// TIA Portal project "消毒机" (V15.1) (continued)
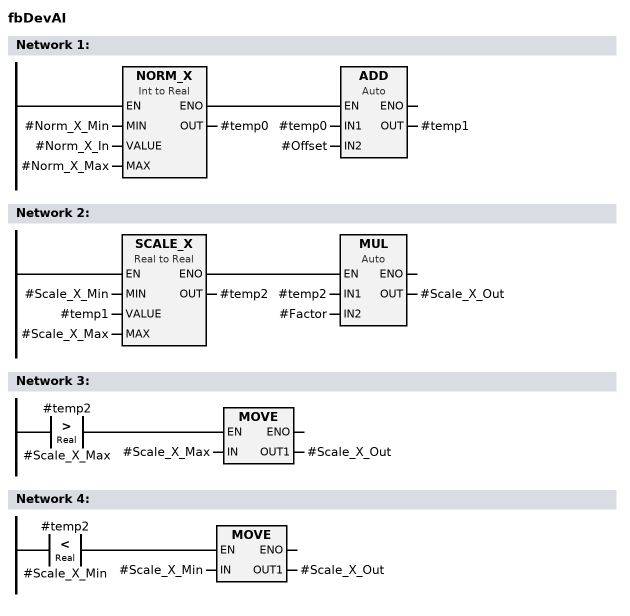
   RUNG wire#powerrail
      { S7_Templates := "[SrcType := Int, DestType := Real]" } Normalize(min := #Norm_X_Min, value := #Norm_X_In, max := #Norm_X_Max, out => #temp0)
      Add(in1 := #temp0, in2 := #Offset, out => #temp1)
   END_RUNG
   // the same network as SCL:
   #temp0 := NORM_X(MIN := #Norm_X_Min, VALUE := #Norm_X_In, MAX := #Norm_X_Max);
   #temp1 := #temp0 + #Offset;
END_REGION

REGION Network 2
   RUNG wire#powerrail
      { S7_Templates := "[SrcType := Real, DestType := Real]" } Scale(min := #Scale_X_Min, value := #temp1, max := #Scale_X_Max, out => #temp2)
      Mul(in1 := #temp2, in2 := #Factor, out => #Scale_X_Out)
   END_RUNG
   // the same network as SCL:
   #temp2 := SCALE_X(MIN := #Scale_X_Min, VALUE := #temp1, MAX := #Scale_X_Max);
   #Scale_X_Out := #temp2 * #Factor;
END_REGION

REGION Network 3
   RUNG wire#powerrail
      { S7_Templates := "SrcType := Real" } GT_Contact(in1 := #temp2, in2 := #Scale_X_Max)
      Move(in := #Scale_X_Max, out1 => #Scale_X_Out)
   END_RUNG
   // the same network as SCL:
   IF #temp2 > #Scale_X_Max THEN #Scale_X_Out := #Scale_X_Max; END_IF;
END_REGION

REGION Network 4
   RUNG wire#powerrail
      { S7_Templates := "SrcType := Real" } LT_Contact(in1 := #temp2, in2 := #Scale_X_Min)
      Move(in := #Scale_X_Min, out1 => #Scale_X_Out)
   END_RUNG
   // the same network as SCL:
   IF #temp2 < #Scale_X_Min THEN #Scale_X_Out := #Scale_X_Min; END_IF;
END_REGION
END_FUNCTION_BLOCK

FUNCTION_BLOCK "fbAI"   // FB102, LAD
{ S7_Optimized_Access := 'TRUE' }
VERSION : 0.1
   VAR
      fbDevAI_Instance : "fbDevAI";
      GET_IM_DATA_Instance : Get_IM_Data;
   END_VAR
   VAR_TEMP
      temp1 : Real;
   END_VAR
BEGIN

REGION Network 1
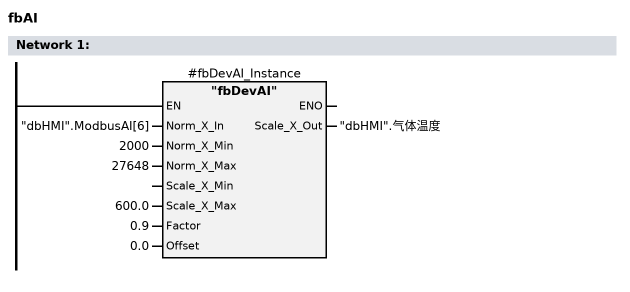
   RUNG wire#powerrail
      #fbDevAI_Instance(Norm_X_In := "dbHMI".ModbusAI[6], Norm_X_Min := 2000, Norm_X_Max := 27648, Scale_X_Min :=, Scale_X_Max := 600.0, Factor := 0.9, Offset := 0.0, Scale_X_Out => "dbHMI".气体温度)
   END_RUNG
   // the same network as SCL:
   #fbDevAI_Instance(Norm_X_In := "dbHMI".ModbusAI[6],   // "fbDevAI"
                     Norm_X_Min := 2000,
                     Norm_X_Max := 27648,
                     Scale_X_Max := 600.0,
                     Factor := 0.9,
                     Offset := 0.0,
                     Scale_X_Out => "dbHMI".气体温度);
END_REGION
END_FUNCTION_BLOCK

FUNCTION_BLOCK "fbSequence"   // FB103, LAD
{ S7_Optimized_Access := 'TRUE' }
VERSION : 0.1
   VAR_INPUT
      Start : Bool;
      Stop : Bool;
      ActUnit : "Unit";
   END_VAR
   VAR_OUTPUT
      ActStepNum : Int;
      OutUnit : "Unit";
   END_VAR
   VAR
      mRuntime_Step : Time;
      sRuntime_Step : Time;
      StepNo : Int;
      "Step" : Array[1..16] of Bool;
      StepDone : Array[1..16] of Bool;
      Next : Bool;
      StepStoped : Array[1..16] of Bool;
      Previos : Bool;
      IEC_Timer_1 : TON_TIME;
      IEC_Timer_2 : TON_TIME;
      IEC_Timer_3 : TON_TIME;
      IEC_Timer_4 : TON_TIME;
      IEC_Timer_5 : TON_TIME;
      IEC_Timer_6 : TON_TIME;
      IEC_Timer_7 : TON_TIME;
      IEC_Timer_8 : TON_TIME;
      IEC_Timer_9 : TON_TIME;
      IEC_Timer_10 : TON_TIME;
      IEC_Timer_11 : TON_TIME;
      IEC_Timer_12 : TON_TIME;
      IEC_Timer_13 : TON_TIME;
      IEC_Timer_14 : TON_TIME;
      IEC_Timer_15 : TON_TIME;
      IEC_Timer_16 : TON_TIME;
      Running : Bool;
      Done : Bool;
      Pls : Array[0..31] of Bool;
      AirCompressor_Step : Array[1..16] of Bool;
      Coolingwater_Step : Array[1..16] of Bool;
      Peristalticpump_Step : Array[1..16] of Bool;
      WepeX_Enable_Step : Array[1..16] of Bool;
      AYV1_Step : Array[1..16] of Bool;
      AYV2_Step : Array[1..16] of Bool;
      BYV1_Step : Array[1..16] of Bool;
      BYV2_Step : Array[1..16] of Bool;
      CYV1_Step : Array[1..16] of Bool;
      CYV2_Step : Array[1..16] of Bool;
      DYV_Step : Array[1..16] of Bool;
      Blower_Step : Array[1..16] of Bool;
   END_VAR
   VAR_TEMP   // added for the SCL form of the ladder/FBD networks
      _w1 : Bool;
   END_VAR
BEGIN

REGION Network 1
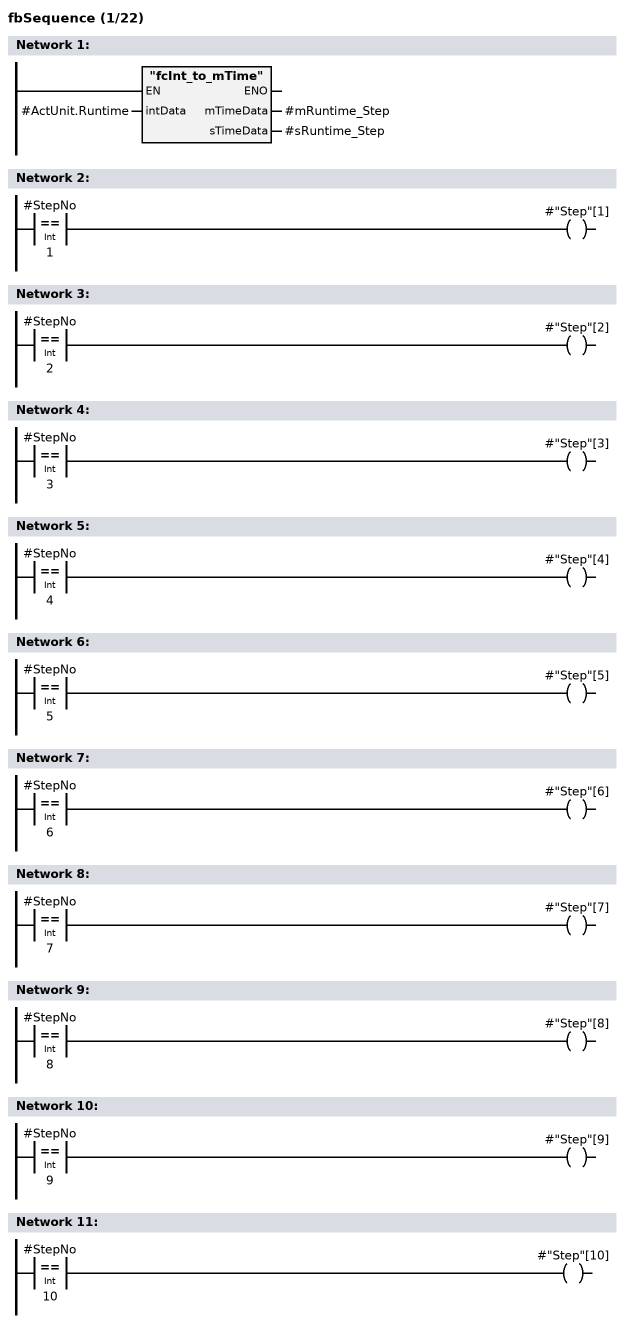
   RUNG wire#powerrail
      "fcInt_to_mTime"(intData := #ActUnit.Runtime, mTimeData => #mRuntime_Step, sTimeData => #sRuntime_Step)
   END_RUNG
   // the same network as SCL:
   "fcInt_to_mTime"(intData := #ActUnit.Runtime, mTimeData => #mRuntime_Step, sTimeData => #sRuntime_Step);
END_REGION

REGION Network 2
   RUNG wire#powerrail
      { S7_Templates := "SrcType := Int" } EQ_Contact(in1 := #StepNo, in2 := 1)
      Coil( #"Step"[1] )
   END_RUNG
   // the same network as SCL:
   #"Step"[1] := #StepNo = 1;
END_REGION

REGION Network 3
   RUNG wire#powerrail
      { S7_Templates := "SrcType := Int" } EQ_Contact(in1 := #StepNo, in2 := 2)
      Coil( #"Step"[2] )
   END_RUNG
   // the same network as SCL:
   #"Step"[2] := #StepNo = 2;
END_REGION

REGION Network 4
   RUNG wire#powerrail
      { S7_Templates := "SrcType := Int" } EQ_Contact(in1 := #StepNo, in2 := 3)
      Coil( #"Step"[3] )
   END_RUNG
   // the same network as SCL:
   #"Step"[3] := #StepNo = 3;
END_REGION

REGION Network 5
   RUNG wire#powerrail
      { S7_Templates := "SrcType := Int" } EQ_Contact(in1 := #StepNo, in2 := 4)
      Coil( #"Step"[4] )
   END_RUNG
   // the same network as SCL:
   #"Step"[4] := #StepNo = 4;
END_REGION

REGION Network 6
   RUNG wire#powerrail
      { S7_Templates := "SrcType := Int" } EQ_Contact(in1 := #StepNo, in2 := 5)
      Coil( #"Step"[5] )
   END_RUNG
   // the same network as SCL:
   #"Step"[5] := #StepNo = 5;
END_REGION

REGION Network 7
   RUNG wire#powerrail
      { S7_Templates := "SrcType := Int" } EQ_Contact(in1 := #StepNo, in2 := 6)
      Coil( #"Step"[6] )
   END_RUNG
   // the same network as SCL:
   #"Step"[6] := #StepNo = 6;
END_REGION

REGION Network 8
   RUNG wire#powerrail
      { S7_Templates := "SrcType := Int" } EQ_Contact(in1 := #StepNo, in2 := 7)
      Coil( #"Step"[7] )
   END_RUNG
   // the same network as SCL:
   #"Step"[7] := #StepNo = 7;
END_REGION

REGION Network 9
   RUNG wire#powerrail
      { S7_Templates := "SrcType := Int" } EQ_Contact(in1 := #StepNo, in2 := 8)
      Coil( #"Step"[8] )
   END_RUNG
   // the same network as SCL:
   #"Step"[8] := #StepNo = 8;
END_REGION

REGION Network 10
   RUNG wire#powerrail
      { S7_Templates := "SrcType := Int" } EQ_Contact(in1 := #StepNo, in2 := 9)
      Coil( #"Step"[9] )
   END_RUNG
   // the same network as SCL:
   #"Step"[9] := #StepNo = 9;
END_REGION

REGION Network 11
   RUNG wire#powerrail
      { S7_Templates := "SrcType := Int" } EQ_Contact(in1 := #StepNo, in2 := 10)
      Coil( #"Step"[10] )
   END_RUNG
   // the same network as SCL:
   #"Step"[10] := #StepNo = 10;
END_REGION

REGION Network 12
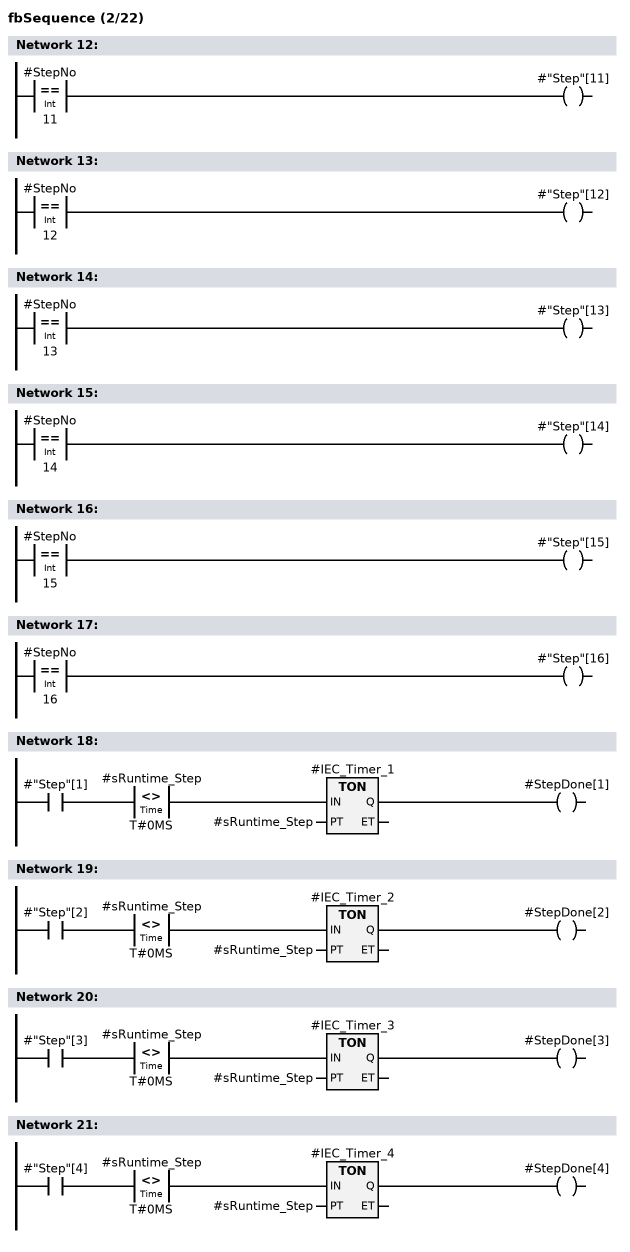
   RUNG wire#powerrail
      { S7_Templates := "SrcType := Int" } EQ_Contact(in1 := #StepNo, in2 := 11)
      Coil( #"Step"[11] )
   END_RUNG
   // the same network as SCL:
   #"Step"[11] := #StepNo = 11;
END_REGION

REGION Network 13
   RUNG wire#powerrail
      { S7_Templates := "SrcType := Int" } EQ_Contact(in1 := #StepNo, in2 := 12)
      Coil( #"Step"[12] )
   END_RUNG
   // the same network as SCL:
   #"Step"[12] := #StepNo = 12;
END_REGION

REGION Network 14
   RUNG wire#powerrail
      { S7_Templates := "SrcType := Int" } EQ_Contact(in1 := #StepNo, in2 := 13)
      Coil( #"Step"[13] )
   END_RUNG
   // the same network as SCL:
   #"Step"[13] := #StepNo = 13;
END_REGION

REGION Network 15
   RUNG wire#powerrail
      { S7_Templates := "SrcType := Int" } EQ_Contact(in1 := #StepNo, in2 := 14)
      Coil( #"Step"[14] )
   END_RUNG
   // the same network as SCL:
   #"Step"[14] := #StepNo = 14;
END_REGION

REGION Network 16
   RUNG wire#powerrail
      { S7_Templates := "SrcType := Int" } EQ_Contact(in1 := #StepNo, in2 := 15)
      Coil( #"Step"[15] )
   END_RUNG
   // the same network as SCL:
   #"Step"[15] := #StepNo = 15;
END_REGION

REGION Network 17
   RUNG wire#powerrail
      { S7_Templates := "SrcType := Int" } EQ_Contact(in1 := #StepNo, in2 := 16)
      Coil( #"Step"[16] )
   END_RUNG
   // the same network as SCL:
   #"Step"[16] := #StepNo = 16;
END_REGION

REGION Network 18
   #IEC_Timer_1(IN := #"Step"[1] AND (#sRuntime_Step <> T#0MS), PT := #sRuntime_Step);   // TON
   #StepDone[1] := #IEC_Timer_1.Q;
END_REGION

REGION Network 19
   #IEC_Timer_2(IN := #"Step"[2] AND (#sRuntime_Step <> T#0MS), PT := #sRuntime_Step);   // TON
   #StepDone[2] := #IEC_Timer_2.Q;
END_REGION

REGION Network 20
   #IEC_Timer_3(IN := #"Step"[3] AND (#sRuntime_Step <> T#0MS), PT := #sRuntime_Step);   // TON
   #StepDone[3] := #IEC_Timer_3.Q;
END_REGION

REGION Network 21
   #IEC_Timer_4(IN := #"Step"[4] AND (#sRuntime_Step <> T#0MS), PT := #sRuntime_Step);   // TON
   #StepDone[4] := #IEC_Timer_4.Q;
END_REGION

REGION Network 22
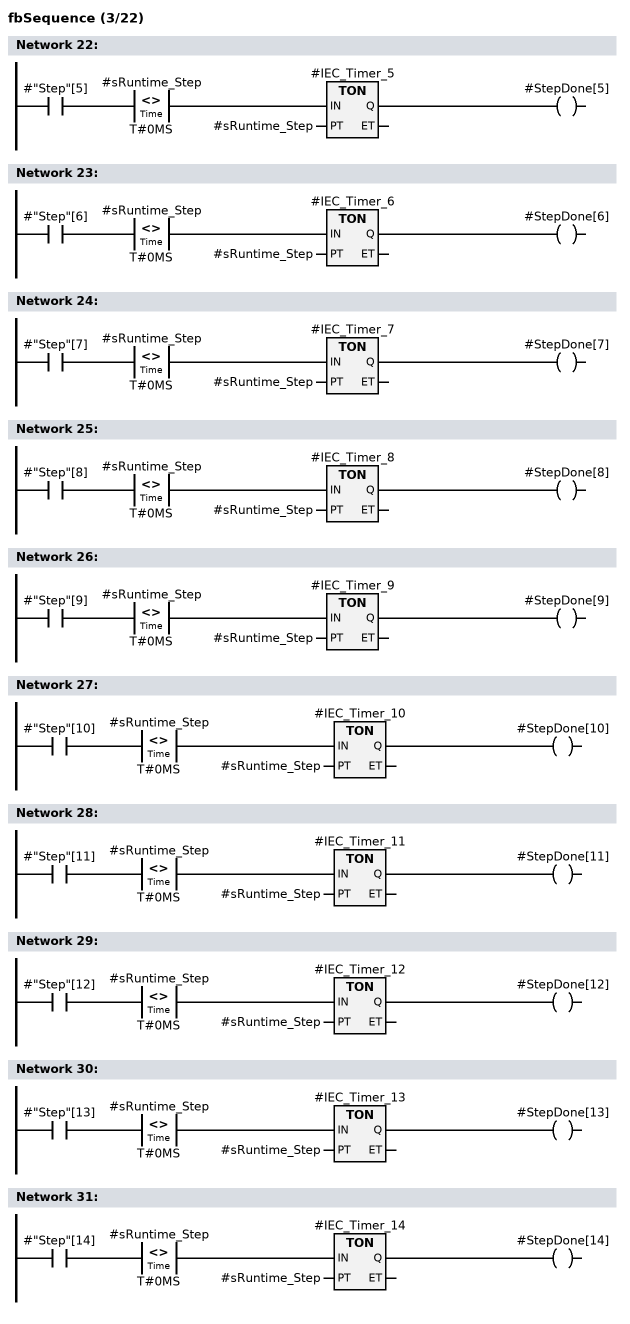
   #IEC_Timer_5(IN := #"Step"[5] AND (#sRuntime_Step <> T#0MS), PT := #sRuntime_Step);   // TON
   #StepDone[5] := #IEC_Timer_5.Q;
END_REGION

REGION Network 23
   #IEC_Timer_6(IN := #"Step"[6] AND (#sRuntime_Step <> T#0MS), PT := #sRuntime_Step);   // TON
   #StepDone[6] := #IEC_Timer_6.Q;
END_REGION

REGION Network 24
   #IEC_Timer_7(IN := #"Step"[7] AND (#sRuntime_Step <> T#0MS), PT := #sRuntime_Step);   // TON
   #StepDone[7] := #IEC_Timer_7.Q;
END_REGION

REGION Network 25
   #IEC_Timer_8(IN := #"Step"[8] AND (#sRuntime_Step <> T#0MS), PT := #sRuntime_Step);   // TON
   #StepDone[8] := #IEC_Timer_8.Q;
END_REGION

REGION Network 26
   #IEC_Timer_9(IN := #"Step"[9] AND (#sRuntime_Step <> T#0MS), PT := #sRuntime_Step);   // TON
   #StepDone[9] := #IEC_Timer_9.Q;
END_REGION

REGION Network 27
   #IEC_Timer_10(IN := #"Step"[10] AND (#sRuntime_Step <> T#0MS), PT := #sRuntime_Step);   // TON
   #StepDone[10] := #IEC_Timer_10.Q;
END_REGION

REGION Network 28
   #IEC_Timer_11(IN := #"Step"[11] AND (#sRuntime_Step <> T#0MS), PT := #sRuntime_Step);   // TON
   #StepDone[11] := #IEC_Timer_11.Q;
END_REGION

REGION Network 29
   #IEC_Timer_12(IN := #"Step"[12] AND (#sRuntime_Step <> T#0MS), PT := #sRuntime_Step);   // TON
   #StepDone[12] := #IEC_Timer_12.Q;
END_REGION

REGION Network 30
   #IEC_Timer_13(IN := #"Step"[13] AND (#sRuntime_Step <> T#0MS), PT := #sRuntime_Step);   // TON
   #StepDone[13] := #IEC_Timer_13.Q;
END_REGION

REGION Network 31
   #IEC_Timer_14(IN := #"Step"[14] AND (#sRuntime_Step <> T#0MS), PT := #sRuntime_Step);   // TON
   #StepDone[14] := #IEC_Timer_14.Q;
END_REGION

REGION Network 32
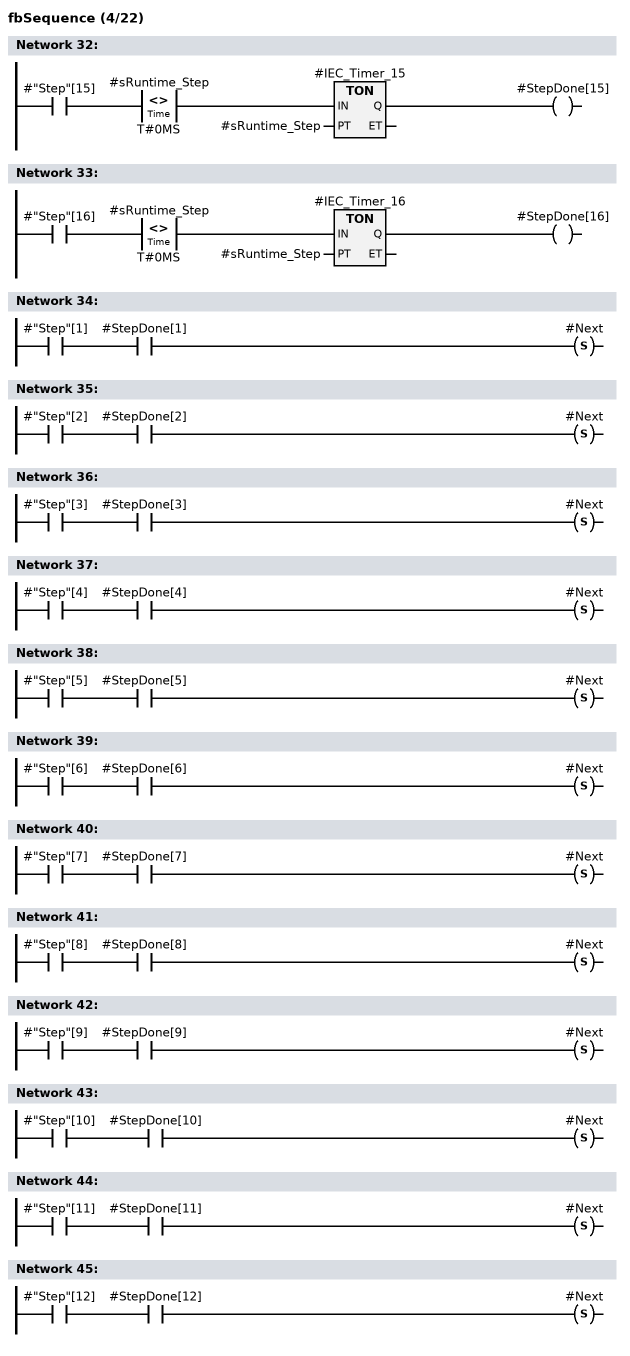
   #IEC_Timer_15(IN := #"Step"[15] AND (#sRuntime_Step <> T#0MS), PT := #sRuntime_Step);   // TON
   #StepDone[15] := #IEC_Timer_15.Q;
END_REGION

REGION Network 33
   #IEC_Timer_16(IN := #"Step"[16] AND (#sRuntime_Step <> T#0MS), PT := #sRuntime_Step);   // TON
   #StepDone[16] := #IEC_Timer_16.Q;
END_REGION

REGION Network 34
   RUNG wire#powerrail
      Contact( #"Step"[1] )
      Contact( #StepDone[1] )
      S_Coil( #Next )
   END_RUNG
   // the same network as SCL:
   IF #"Step"[1] AND #StepDone[1] THEN #Next := TRUE; END_IF;
END_REGION

REGION Network 35
   RUNG wire#powerrail
      Contact( #"Step"[2] )
      Contact( #StepDone[2] )
      S_Coil( #Next )
   END_RUNG
   // the same network as SCL:
   IF #"Step"[2] AND #StepDone[2] THEN #Next := TRUE; END_IF;
END_REGION

REGION Network 36
   RUNG wire#powerrail
      Contact( #"Step"[3] )
      Contact( #StepDone[3] )
      S_Coil( #Next )
   END_RUNG
   // the same network as SCL:
   IF #"Step"[3] AND #StepDone[3] THEN #Next := TRUE; END_IF;
END_REGION

REGION Network 37
   RUNG wire#powerrail
      Contact( #"Step"[4] )
      Contact( #StepDone[4] )
      S_Coil( #Next )
   END_RUNG
   // the same network as SCL:
   IF #"Step"[4] AND #StepDone[4] THEN #Next := TRUE; END_IF;
END_REGION

REGION Network 38
   RUNG wire#powerrail
      Contact( #"Step"[5] )
      Contact( #StepDone[5] )
      S_Coil( #Next )
   END_RUNG
   // the same network as SCL:
   IF #"Step"[5] AND #StepDone[5] THEN #Next := TRUE; END_IF;
END_REGION

REGION Network 39
   RUNG wire#powerrail
      Contact( #"Step"[6] )
      Contact( #StepDone[6] )
      S_Coil( #Next )
   END_RUNG
   // the same network as SCL:
   IF #"Step"[6] AND #StepDone[6] THEN #Next := TRUE; END_IF;
END_REGION

REGION Network 40
   RUNG wire#powerrail
      Contact( #"Step"[7] )
      Contact( #StepDone[7] )
      S_Coil( #Next )
   END_RUNG
   // the same network as SCL:
   IF #"Step"[7] AND #StepDone[7] THEN #Next := TRUE; END_IF;
END_REGION

REGION Network 41
   RUNG wire#powerrail
      Contact( #"Step"[8] )
      Contact( #StepDone[8] )
      S_Coil( #Next )
   END_RUNG
   // the same network as SCL:
   IF #"Step"[8] AND #StepDone[8] THEN #Next := TRUE; END_IF;
END_REGION

REGION Network 42
   RUNG wire#powerrail
      Contact( #"Step"[9] )
      Contact( #StepDone[9] )
      S_Coil( #Next )
   END_RUNG
   // the same network as SCL:
   IF #"Step"[9] AND #StepDone[9] THEN #Next := TRUE; END_IF;
END_REGION

REGION Network 43
   RUNG wire#powerrail
      Contact( #"Step"[10] )
      Contact( #StepDone[10] )
      S_Coil( #Next )
   END_RUNG
   // the same network as SCL:
   IF #"Step"[10] AND #StepDone[10] THEN #Next := TRUE; END_IF;
END_REGION

REGION Network 44
   RUNG wire#powerrail
      Contact( #"Step"[11] )
      Contact( #StepDone[11] )
      S_Coil( #Next )
   END_RUNG
   // the same network as SCL:
   IF #"Step"[11] AND #StepDone[11] THEN #Next := TRUE; END_IF;
END_REGION

REGION Network 45
   RUNG wire#powerrail
      Contact( #"Step"[12] )
      Contact( #StepDone[12] )
      S_Coil( #Next )
   END_RUNG
   // the same network as SCL:
   IF #"Step"[12] AND #StepDone[12] THEN #Next := TRUE; END_IF;
END_REGION

REGION Network 46
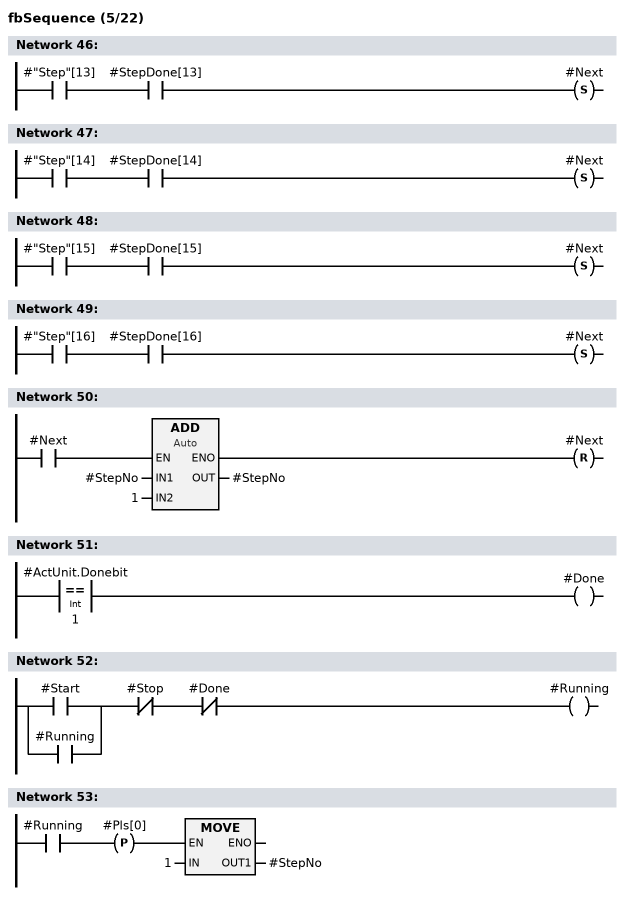
   RUNG wire#powerrail
      Contact( #"Step"[13] )
      Contact( #StepDone[13] )
      S_Coil( #Next )
   END_RUNG
   // the same network as SCL:
   IF #"Step"[13] AND #StepDone[13] THEN #Next := TRUE; END_IF;
END_REGION

REGION Network 47
   RUNG wire#powerrail
      Contact( #"Step"[14] )
      Contact( #StepDone[14] )
      S_Coil( #Next )
   END_RUNG
   // the same network as SCL:
   IF #"Step"[14] AND #StepDone[14] THEN #Next := TRUE; END_IF;
END_REGION

REGION Network 48
   RUNG wire#powerrail
      Contact( #"Step"[15] )
      Contact( #StepDone[15] )
      S_Coil( #Next )
   END_RUNG
   // the same network as SCL:
   IF #"Step"[15] AND #StepDone[15] THEN #Next := TRUE; END_IF;
END_REGION

REGION Network 49
   RUNG wire#powerrail
      Contact( #"Step"[16] )
      Contact( #StepDone[16] )
      S_Coil( #Next )
   END_RUNG
   // the same network as SCL:
   IF #"Step"[16] AND #StepDone[16] THEN #Next := TRUE; END_IF;
END_REGION

REGION Network 50
   RUNG wire#powerrail
      Contact( #Next )
      Add(in1 := #StepNo, in2 := 1, out => #StepNo)
      R_Coil( #Next )
   END_RUNG
   // the same network as SCL:
   IF #Next THEN
       #StepNo := #StepNo + 1;
       #Next := FALSE;
   END_IF;
END_REGION

REGION Network 51
   RUNG wire#powerrail
      { S7_Templates := "SrcType := Int" } EQ_Contact(in1 := #ActUnit.Donebit, in2 := 1)
      Coil( #Done )
   END_RUNG
   // the same network as SCL:
   #Done := #ActUnit.Donebit = 1;
END_REGION

REGION Network 52
   RUNG wire#powerrail
      Contact( #Start )
      wire#w1
      I_Contact( #Stop )
      I_Contact( #Done )
      Coil( #Running )
   END_RUNG
   RUNG wire#powerrail
      Contact( #Running )
   END_RUNG wire#w1
   // the same network as SCL:
   #Running := (#Start OR #Running) AND NOT #Stop AND NOT #Done;
END_REGION

REGION Network 53
   RUNG wire#powerrail
      Contact( #Running )
      P_Trig( #Pls[0] )
      Move(in := 1, out1 => #StepNo)
   END_RUNG
   // the same network as SCL:
   #_w1 := #Running AND NOT #Pls[0];   // rising edge
   #Pls[0] := #Running;
   IF #_w1 THEN #StepNo := 1; END_IF;
END_REGION

REGION Network 54
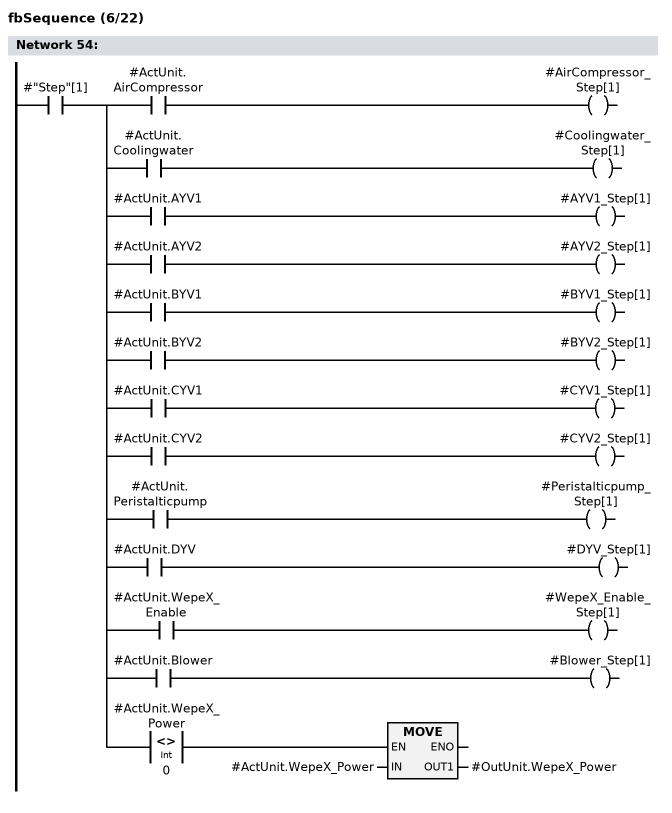
   RUNG wire#powerrail
      Contact( #"Step"[1] )
      wire#w1
      Contact( #ActUnit.AirCompressor )
      Coil( #AirCompressor_Step[1] )
   END_RUNG
   RUNG wire#w1
      Contact( #ActUnit.Coolingwater )
      Coil( #Coolingwater_Step[1] )
   END_RUNG
   RUNG wire#w1
      Contact( #ActUnit.AYV1 )
      Coil( #AYV1_Step[1] )
   END_RUNG
   RUNG wire#w1
      Contact( #ActUnit.AYV2 )
      Coil( #AYV2_Step[1] )
   END_RUNG
   RUNG wire#w1
      Contact( #ActUnit.BYV1 )
      Coil( #BYV1_Step[1] )
   END_RUNG
   RUNG wire#w1
      Contact( #ActUnit.BYV2 )
      Coil( #BYV2_Step[1] )
   END_RUNG
   RUNG wire#w1
      Contact( #ActUnit.CYV1 )
      Coil( #CYV1_Step[1] )
   END_RUNG
   RUNG wire#w1
      Contact( #ActUnit.CYV2 )
      Coil( #CYV2_Step[1] )
   END_RUNG
   RUNG wire#w1
      Contact( #ActUnit.Peristalticpump )
      Coil( #Peristalticpump_Step[1] )
   END_RUNG
   RUNG wire#w1
      Contact( #ActUnit.DYV )
      Coil( #DYV_Step[1] )
   END_RUNG
   RUNG wire#w1
      Contact( #ActUnit.WepeX_Enable )
      Coil( #WepeX_Enable_Step[1] )
   END_RUNG
   RUNG wire#w1
      Contact( #ActUnit.Blower )
      Coil( #Blower_Step[1] )
   END_RUNG
   RUNG wire#w1
      { S7_Templates := "SrcType := Int" } NE_Contact(in1 := #ActUnit.WepeX_Power, in2 := 0)
      Move(in := #ActUnit.WepeX_Power, out1 => #OutUnit.WepeX_Power)
   END_RUNG
   // the same network as SCL:
   #AirCompressor_Step[1] := #"Step"[1] AND #ActUnit.AirCompressor;
   #Coolingwater_Step[1] := #"Step"[1] AND #ActUnit.Coolingwater;
   #AYV1_Step[1] := #"Step"[1] AND #ActUnit.AYV1;
   #AYV2_Step[1] := #"Step"[1] AND #ActUnit.AYV2;
   #BYV1_Step[1] := #"Step"[1] AND #ActUnit.BYV1;
   #BYV2_Step[1] := #"Step"[1] AND #ActUnit.BYV2;
   #CYV1_Step[1] := #"Step"[1] AND #ActUnit.CYV1;
   #CYV2_Step[1] := #"Step"[1] AND #ActUnit.CYV2;
   #Peristalticpump_Step[1] := #"Step"[1] AND #ActUnit.Peristalticpump;
   #DYV_Step[1] := #"Step"[1] AND #ActUnit.DYV;
   #WepeX_Enable_Step[1] := #"Step"[1] AND #ActUnit.WepeX_Enable;
   #Blower_Step[1] := #"Step"[1] AND #ActUnit.Blower;
   IF #"Step"[1] AND (#ActUnit.WepeX_Power <> 0) THEN #OutUnit.WepeX_Power := #ActUnit.WepeX_Power; END_IF;
END_REGION

REGION Network 55
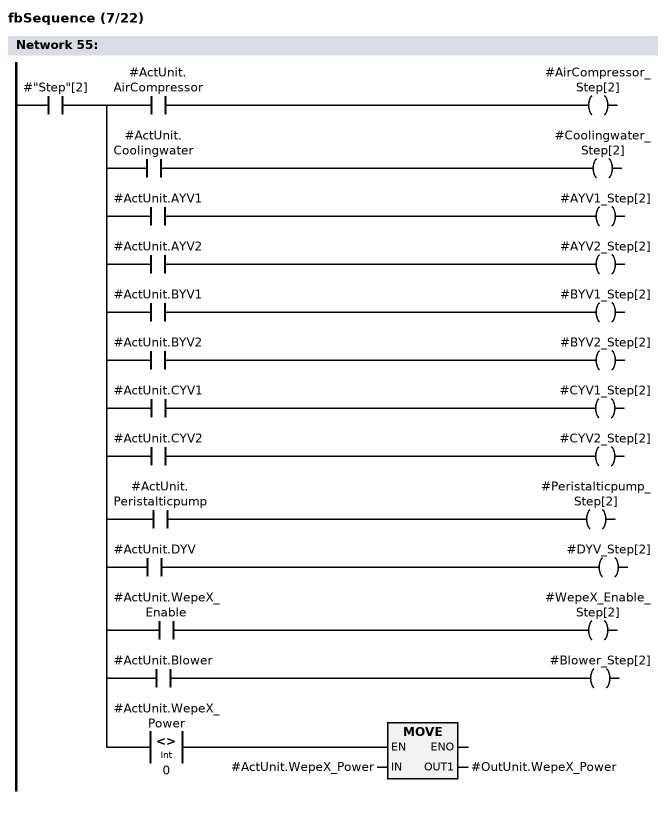
   RUNG wire#powerrail
      Contact( #"Step"[2] )
      wire#w1
      Contact( #ActUnit.AirCompressor )
      Coil( #AirCompressor_Step[2] )
   END_RUNG
   RUNG wire#w1
      Contact( #ActUnit.Coolingwater )
      Coil( #Coolingwater_Step[2] )
   END_RUNG
   RUNG wire#w1
      Contact( #ActUnit.AYV1 )
      Coil( #AYV1_Step[2] )
   END_RUNG
   RUNG wire#w1
      Contact( #ActUnit.AYV2 )
      Coil( #AYV2_Step[2] )
   END_RUNG
   RUNG wire#w1
      Contact( #ActUnit.BYV1 )
      Coil( #BYV1_Step[2] )
   END_RUNG
   RUNG wire#w1
      Contact( #ActUnit.BYV2 )
      Coil( #BYV2_Step[2] )
   END_RUNG
   RUNG wire#w1
      Contact( #ActUnit.CYV1 )
      Coil( #CYV1_Step[2] )
   END_RUNG
   RUNG wire#w1
      Contact( #ActUnit.CYV2 )
      Coil( #CYV2_Step[2] )
   END_RUNG
   RUNG wire#w1
      Contact( #ActUnit.Peristalticpump )
      Coil( #Peristalticpump_Step[2] )
   END_RUNG
   RUNG wire#w1
      Contact( #ActUnit.DYV )
      Coil( #DYV_Step[2] )
   END_RUNG
   RUNG wire#w1
      Contact( #ActUnit.WepeX_Enable )
      Coil( #WepeX_Enable_Step[2] )
   END_RUNG
   RUNG wire#w1
      Contact( #ActUnit.Blower )
      Coil( #Blower_Step[2] )
   END_RUNG
   RUNG wire#w1
      { S7_Templates := "SrcType := Int" } NE_Contact(in1 := #ActUnit.WepeX_Power, in2 := 0)
      Move(in := #ActUnit.WepeX_Power, out1 => #OutUnit.WepeX_Power)
   END_RUNG
   // the same network as SCL:
   #AirCompressor_Step[2] := #"Step"[2] AND #ActUnit.AirCompressor;
   #Coolingwater_Step[2] := #"Step"[2] AND #ActUnit.Coolingwater;
   #AYV1_Step[2] := #"Step"[2] AND #ActUnit.AYV1;
   #AYV2_Step[2] := #"Step"[2] AND #ActUnit.AYV2;
   #BYV1_Step[2] := #"Step"[2] AND #ActUnit.BYV1;
   #BYV2_Step[2] := #"Step"[2] AND #ActUnit.BYV2;
   #CYV1_Step[2] := #"Step"[2] AND #ActUnit.CYV1;
   #CYV2_Step[2] := #"Step"[2] AND #ActUnit.CYV2;
   #Peristalticpump_Step[2] := #"Step"[2] AND #ActUnit.Peristalticpump;
   #DYV_Step[2] := #"Step"[2] AND #ActUnit.DYV;
   #WepeX_Enable_Step[2] := #"Step"[2] AND #ActUnit.WepeX_Enable;
   #Blower_Step[2] := #"Step"[2] AND #ActUnit.Blower;
   IF #"Step"[2] AND (#ActUnit.WepeX_Power <> 0) THEN #OutUnit.WepeX_Power := #ActUnit.WepeX_Power; END_IF;
END_REGION

REGION Network 56